REGION Network 8: UnHold Command - controlled by Category Alarm 7
   RUNG wire#powerrail
      Contact( "PackML".Sts.State.Held )
      I_Contact( "UN".Alarm.sts_Category_7_NotLatched )
      Coil( "UN".PackML_Sts_Alarm.cmd_UnHold )
   END_RUNG
   // the same network as SCL:
   "UN".PackML_Sts_Alarm.cmd_UnHold := "PackML".Sts.State.Held AND NOT "UN".Alarm.sts_Category_7_NotLatched;
END_REGION

REGION Network 9: Suspend Command - controlled by Category Alarm 8 or 9
   RUNG wire#powerrail
      Contact( "UN".Alarm.sts_Category_8_NotLatched )
      wire#w1
      Coil( "UN".PackML_Sts_Alarm.cmd_Suspend )
   END_RUNG
   RUNG wire#powerrail
      Contact( "UN".Alarm.sts_Category_9_NotLatched )
   END_RUNG wire#w1
   // the same network as SCL:
   "UN".PackML_Sts_Alarm.cmd_Suspend := "UN".Alarm.sts_Category_8_NotLatched OR "UN".Alarm.sts_Category_9_NotLatched;
END_REGION

REGION Network 10: UnSuspend Command - controlled by clearedCategory Alarm 8 or 9
   RUNG wire#powerrail
      Contact( "PackML".Sts.State.Suspended )
      I_Contact( "UN".Alarm.sts_Category_8_NotLatched )
      I_Contact( "UN".Alarm.sts_Category_9_NotLatched )
      Coil( "UN".PackML_Sts_Alarm.cmd_UnSuspend )
   END_RUNG
   // the same network as SCL:
   "UN".PackML_Sts_Alarm.cmd_UnSuspend := "PackML".Sts.State.Suspended AND NOT "UN".Alarm.sts_Category_8_NotLatched AND NOT "UN".Alarm.sts_Category_9_NotLatched;
END_REGION

REGION Network 11: Clearing SC Command - controlled by clearedCategory Alarm 0 or 1
   RUNG wire#powerrail
      Contact( "PackML".Sts.State.Clearing )
      I_Contact( "UN".Alarm.sts_Category_0_Latched )
      I_Contact( "UN".Alarm.sts_Category_1_Latched )
      Coil( "UN".PackML_Sts_Alarm.sts_Clearing_SC )
   END_RUNG
   // the same network as SCL:
   "UN".PackML_Sts_Alarm.sts_Clearing_SC := "PackML".Sts.State.Clearing AND NOT "UN".Alarm.sts_Category_0_Latched AND NOT "UN".Alarm.sts_Category_1_Latched;
END_REGION

REGION Network 12: Resetting S Command - controlled by clearedCategory Alarm 0-4
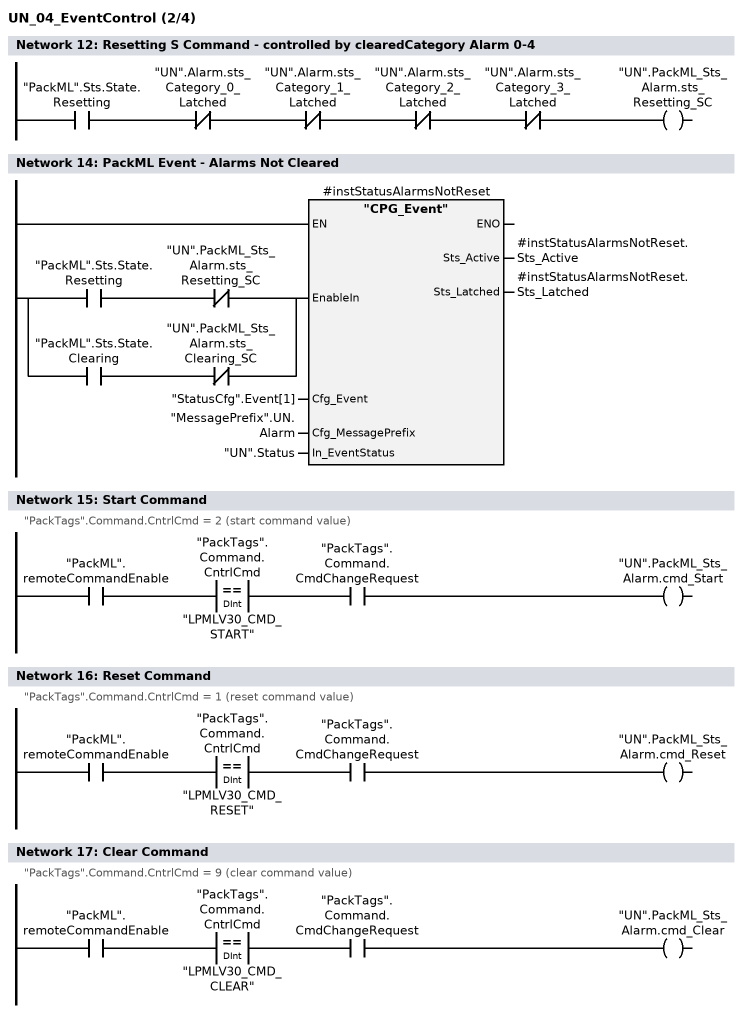
   RUNG wire#powerrail
      Contact( "PackML".Sts.State.Resetting )
      I_Contact( "UN".Alarm.sts_Category_0_Latched )
      I_Contact( "UN".Alarm.sts_Category_1_Latched )
      I_Contact( "UN".Alarm.sts_Category_2_Latched )
      I_Contact( "UN".Alarm.sts_Category_3_Latched )
      Coil( "UN".PackML_Sts_Alarm.sts_Resetting_SC )
   END_RUNG
   // the same network as SCL:
   "UN".PackML_Sts_Alarm.sts_Resetting_SC := "PackML".Sts.State.Resetting AND NOT "UN".Alarm.sts_Category_0_Latched AND NOT "UN".Alarm.sts_Category_1_Latched AND NOT "UN".Alarm.sts_Category_2_Latched AND NOT "UN".Alarm.sts_Category_3_Latched;
END_REGION

REGION Network 13: PackML Event -
END_REGION

REGION Network 14: PackML Event - Alarms Not Cleared
   RUNG wire#powerrail
      #instStatusAlarmsNotReset(EnableIn := wire#w1, Cfg_Event := "StatusCfg".Event[1], Cfg_MessagePrefix := "MessagePrefix".UN.Alarm, In_EventStatus := "UN".Status, Sts_Active => #instStatusAlarmsNotReset.Sts_Active, Sts_Latched => #instStatusAlarmsNotReset.Sts_Latched)
   END_RUNG
   RUNG wire#powerrail
      Contact( "PackML".Sts.State.Resetting )
      I_Contact( "UN".PackML_Sts_Alarm.sts_Resetting_SC )
   END_RUNG wire#w1
   RUNG wire#powerrail
      Contact( "PackML".Sts.State.Clearing )
      I_Contact( "UN".PackML_Sts_Alarm.sts_Clearing_SC )
   END_RUNG wire#w1
   // the same network as SCL:
   #instStatusAlarmsNotReset(EnableIn := ("PackML".Sts.State.Resetting AND NOT "UN".PackML_Sts_Alarm.sts_Resetting_SC) OR ("PackML".Sts.State.Clearing AND NOT "UN".PackML_Sts_Alarm.sts_Clearing_SC),   // "CPG_Event"
                           Cfg_Event := "StatusCfg".Event[1],
                           Cfg_MessagePrefix := "MessagePrefix".UN.Alarm,
                           In_EventStatus := "UN".Status,
                           Sts_Active => #instStatusAlarmsNotReset.Sts_Active,
                           Sts_Latched => #instStatusAlarmsNotReset.Sts_Latched);
END_REGION

REGION Network 15: Start Command
   // "PackTags".Command.CntrlCmd = 2 (start command value)
   RUNG wire#powerrail
      Contact( "PackML".remoteCommandEnable )
      { S7_Templates := "SrcType := DInt" } EQ_Contact(in1 := "PackTags".Command.CntrlCmd, in2 := "LPMLV30_CMD_START")
      Contact( "PackTags".Command.CmdChangeRequest )
      Coil( "UN".PackML_Sts_Alarm.cmd_Start )
   END_RUNG
   // the same network as SCL:
   "UN".PackML_Sts_Alarm.cmd_Start := "PackML".remoteCommandEnable AND ("PackTags".Command.CntrlCmd = "LPMLV30_CMD_START") AND "PackTags".Command.CmdChangeRequest;
END_REGION

REGION Network 16: Reset Command
   // "PackTags".Command.CntrlCmd = 1 (reset command value)
   RUNG wire#powerrail
      Contact( "PackML".remoteCommandEnable )
      { S7_Templates := "SrcType := DInt" } EQ_Contact(in1 := "PackTags".Command.CntrlCmd, in2 := "LPMLV30_CMD_RESET")
      Contact( "PackTags".Command.CmdChangeRequest )
      Coil( "UN".PackML_Sts_Alarm.cmd_Reset )
   END_RUNG
   // the same network as SCL:
   "UN".PackML_Sts_Alarm.cmd_Reset := "PackML".remoteCommandEnable AND ("PackTags".Command.CntrlCmd = "LPMLV30_CMD_RESET") AND "PackTags".Command.CmdChangeRequest;
END_REGION

REGION Network 17: Clear Command
   // "PackTags".Command.CntrlCmd = 9 (clear command value)
   RUNG wire#powerrail
      Contact( "PackML".remoteCommandEnable )
      { S7_Templates := "SrcType := DInt" } EQ_Contact(in1 := "PackTags".Command.CntrlCmd, in2 := "LPMLV30_CMD_CLEAR")
      Contact( "PackTags".Command.CmdChangeRequest )
      Coil( "UN".PackML_Sts_Alarm.cmd_Clear )
   END_RUNG
   // the same network as SCL:
   "UN".PackML_Sts_Alarm.cmd_Clear := "PackML".remoteCommandEnable AND ("PackTags".Command.CntrlCmd = "LPMLV30_CMD_CLEAR") AND "PackTags".Command.CmdChangeRequest;
END_REGION

REGION Network 18: *** EVENT CONTROL MANAGERS ***
END_REGION

REGION Network 19: Reset Command - for all event managers
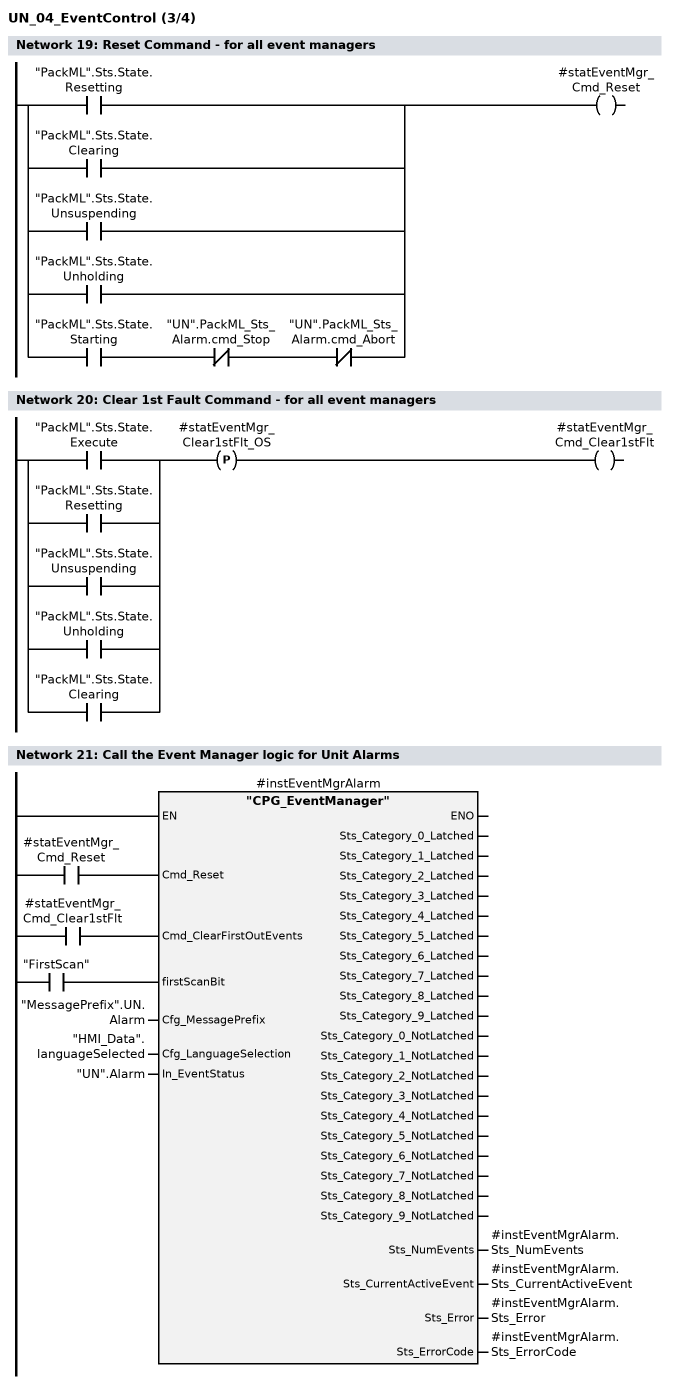
   RUNG wire#powerrail
      Contact( "PackML".Sts.State.Resetting )
      wire#w1
      Coil( #statEventMgr_Cmd_Reset )
   END_RUNG
   RUNG wire#powerrail
      Contact( "PackML".Sts.State.Clearing )
   END_RUNG wire#w1
   RUNG wire#powerrail
      Contact( "PackML".Sts.State.Unsuspending )
   END_RUNG wire#w1
   RUNG wire#powerrail
      Contact( "PackML".Sts.State.Unholding )
   END_RUNG wire#w1
   RUNG wire#powerrail
      Contact( "PackML".Sts.State.Starting )
      I_Contact( "UN".PackML_Sts_Alarm.cmd_Stop )
      I_Contact( "UN".PackML_Sts_Alarm.cmd_Abort )
   END_RUNG wire#w1
   // the same network as SCL:
   #statEventMgr_Cmd_Reset := "PackML".Sts.State.Resetting OR "PackML".Sts.State.Clearing OR "PackML".Sts.State.Unsuspending OR "PackML".Sts.State.Unholding OR ("PackML".Sts.State.Starting AND NOT "UN".PackML_Sts_Alarm.cmd_Stop AND NOT "UN".PackML_Sts_Alarm.cmd_Abort);
END_REGION

REGION Network 20: Clear 1st Fault Command - for all event managers
   RUNG wire#powerrail
      Contact( "PackML".Sts.State.Execute )
      wire#w1
      P_Trig( #statEventMgr_Clear1stFlt_OS )
      Coil( #statEventMgr_Cmd_Clear1stFlt )
   END_RUNG
   RUNG wire#powerrail
      Contact( "PackML".Sts.State.Resetting )
   END_RUNG wire#w1
   RUNG wire#powerrail
      Contact( "PackML".Sts.State.Unsuspending )
   END_RUNG wire#w1
   RUNG wire#powerrail
      Contact( "PackML".Sts.State.Unholding )
   END_RUNG wire#w1
   RUNG wire#powerrail
      Contact( "PackML".Sts.State.Clearing )
   END_RUNG wire#w1
   // the same network as SCL:
   #_w1 := "PackML".Sts.State.Execute OR "PackML".Sts.State.Resetting OR "PackML".Sts.State.Unsuspending OR "PackML".Sts.State.Unholding OR "PackML".Sts.State.Clearing;
   #_w2 := #_w1 AND NOT #statEventMgr_Clear1stFlt_OS;   // rising edge
   #statEventMgr_Clear1stFlt_OS := #_w1;
   #statEventMgr_Cmd_Clear1stFlt := #_w2;
END_REGION

REGION Network 21: Call the Event Manager logic for Unit Alarms
   RUNG wire#powerrail
      #instEventMgrAlarm(Cmd_Reset := wire#w1, Cmd_ClearFirstOutEvents := wire#w2, firstScanBit := wire#w3, Cfg_MessagePrefix := "MessagePrefix".UN.Alarm, Cfg_LanguageSelection := "HMI_Data".languageSelected, In_EventStatus := "UN".Alarm, Sts_Category_0_Latched =>, Sts_Category_1_Latched =>, Sts_Category_2_Latched =>, Sts_Category_3_Latched =>, Sts_Category_4_Latched =>, Sts_Category_5_Latched =>, Sts_Category_6_Latched =>, Sts_Category_7_Latched =>, Sts_Category_8_Latched =>, Sts_Category_9_Latched =>, Sts_Category_0_NotLatched =>, Sts_Category_1_NotLatched =>, Sts_Category_2_NotLatched =>, Sts_Category_3_NotLatched =>, Sts_Category_4_NotLatched =>, Sts_Category_5_NotLatched =>, Sts_Category_6_NotLatched =>, Sts_Category_7_NotLatched =>, Sts_Category_8_NotLatched =>, Sts_Category_9_NotLatched =>, Sts_NumEvents => #instEventMgrAlarm.Sts_NumEvents, Sts_CurrentActiveEvent => #instEventMgrAlarm.Sts_CurrentActiveEvent, Sts_Error => #instEventMgrAlarm.Sts_Error, Sts_ErrorCode => #instEventMgrAlarm.Sts_ErrorCode)
   END_RUNG
   RUNG wire#powerrail
      Contact( #statEventMgr_Cmd_Reset )
   END_RUNG wire#w1
   RUNG wire#powerrail
      Contact( #statEventMgr_Cmd_Clear1stFlt )
   END_RUNG wire#w2
   RUNG wire#powerrail
      Contact( "FirstScan" )
   END_RUNG wire#w3
   // the same network as SCL:
   #instEventMgrAlarm(Cmd_Reset := #statEventMgr_Cmd_Reset,   // "CPG_EventManager"
                      Cmd_ClearFirstOutEvents := #statEventMgr_Cmd_Clear1stFlt,
                      firstScanBit := "FirstScan",
                      Cfg_MessagePrefix := "MessagePrefix".UN.Alarm,
                      Cfg_LanguageSelection := "HMI_Data".languageSelected,
                      In_EventStatus := "UN".Alarm,
                      Sts_NumEvents => #instEventMgrAlarm.Sts_NumEvents,
                      Sts_CurrentActiveEvent => #instEventMgrAlarm.Sts_CurrentActiveEvent,
                      Sts_Error => #instEventMgrAlarm.Sts_Error,
                      Sts_ErrorCode => #instEventMgrAlarm.Sts_ErrorCode);
END_REGION

REGION Network 22: Call the Event Manager logic for Unit Warnings
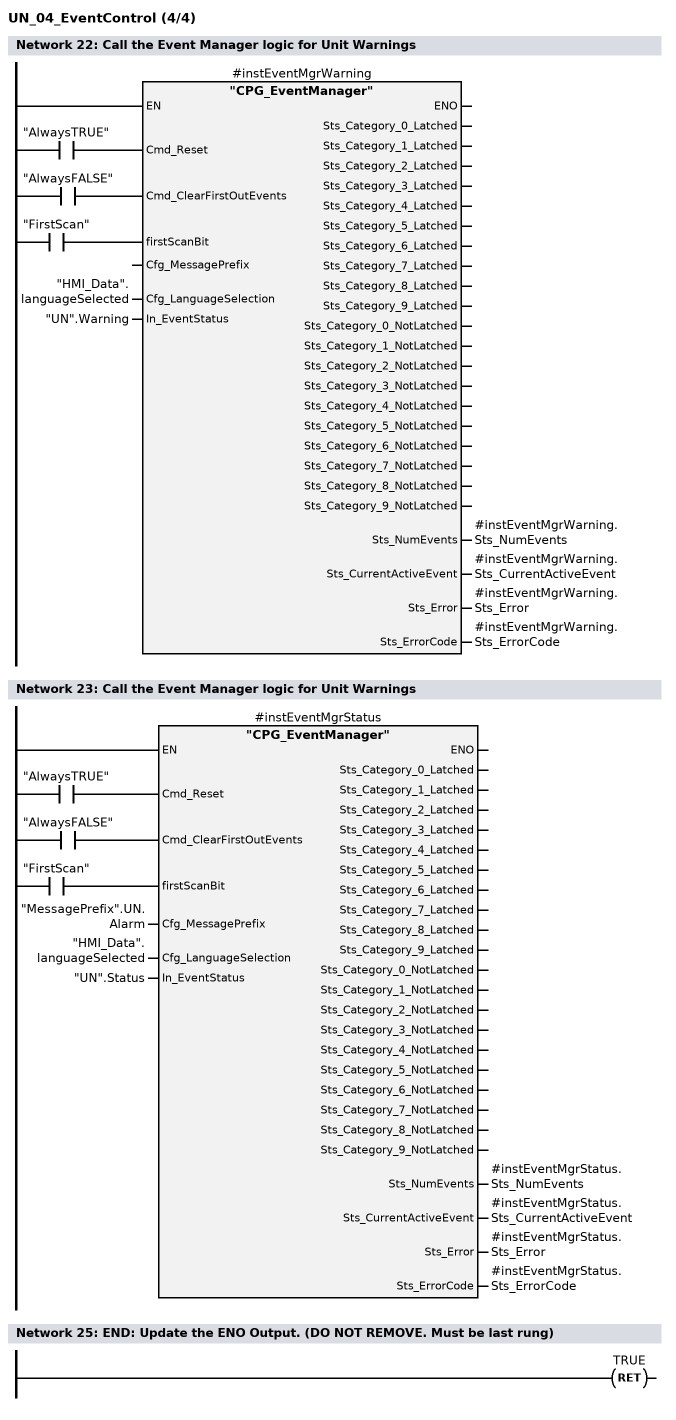
   RUNG wire#powerrail
      #instEventMgrWarning(Cmd_Reset := wire#w1, Cmd_ClearFirstOutEvents := wire#w2, firstScanBit := wire#w3, Cfg_MessagePrefix :=, Cfg_LanguageSelection := "HMI_Data".languageSelected, In_EventStatus := "UN".Warning, Sts_Category_0_Latched =>, Sts_Category_1_Latched =>, Sts_Category_2_Latched =>, Sts_Category_3_Latched =>, Sts_Category_4_Latched =>, Sts_Category_5_Latched =>, Sts_Category_6_Latched =>, Sts_Category_7_Latched =>, Sts_Category_8_Latched =>, Sts_Category_9_Latched =>, Sts_Category_0_NotLatched =>, Sts_Category_1_NotLatched =>, Sts_Category_2_NotLatched =>, Sts_Category_3_NotLatched =>, Sts_Category_4_NotLatched =>, Sts_Category_5_NotLatched =>, Sts_Category_6_NotLatched =>, Sts_Category_7_NotLatched =>, Sts_Category_8_NotLatched =>, Sts_Category_9_NotLatched =>, Sts_NumEvents => #instEventMgrWarning.Sts_NumEvents, Sts_CurrentActiveEvent => #instEventMgrWarning.Sts_CurrentActiveEvent, Sts_Error => #instEventMgrWarning.Sts_Error, Sts_ErrorCode => #instEventMgrWarning.Sts_ErrorCode)
   END_RUNG
   RUNG wire#powerrail
      Contact( "AlwaysTRUE" )
   END_RUNG wire#w1
   RUNG wire#powerrail
      Contact( "AlwaysFALSE" )
   END_RUNG wire#w2
   RUNG wire#powerrail
      Contact( "FirstScan" )
   END_RUNG wire#w3
   // the same network as SCL:
   #instEventMgrWarning(Cmd_Reset := "AlwaysTRUE",   // "CPG_EventManager"
                        Cmd_ClearFirstOutEvents := "AlwaysFALSE",
                        firstScanBit := "FirstScan",
                        Cfg_LanguageSelection := "HMI_Data".languageSelected,
                        In_EventStatus := "UN".Warning,
                        Sts_NumEvents => #instEventMgrWarning.Sts_NumEvents,
                        Sts_CurrentActiveEvent => #instEventMgrWarning.Sts_CurrentActiveEvent,
                        Sts_Error => #instEventMgrWarning.Sts_Error,
                        Sts_ErrorCode => #instEventMgrWarning.Sts_ErrorCode);
END_REGION

REGION Network 23: Call the Event Manager logic for Unit Warnings
   RUNG wire#powerrail
      #instEventMgrStatus(Cmd_Reset := wire#w1, Cmd_ClearFirstOutEvents := wire#w2, firstScanBit := wire#w3, Cfg_MessagePrefix := "MessagePrefix".UN.Alarm, Cfg_LanguageSelection := "HMI_Data".languageSelected, In_EventStatus := "UN".Status, Sts_Category_0_Latched =>, Sts_Category_1_Latched =>, Sts_Category_2_Latched =>, Sts_Category_3_Latched =>, Sts_Category_4_Latched =>, Sts_Category_5_Latched =>, Sts_Category_6_Latched =>, Sts_Category_7_Latched =>, Sts_Category_8_Latched =>, Sts_Category_9_Latched =>, Sts_Category_0_NotLatched =>, Sts_Category_1_NotLatched =>, Sts_Category_2_NotLatched =>, Sts_Category_3_NotLatched =>, Sts_Category_4_NotLatched =>, Sts_Category_5_NotLatched =>, Sts_Category_6_NotLatched =>, Sts_Category_7_NotLatched =>, Sts_Category_8_NotLatched =>, Sts_Category_9_NotLatched =>, Sts_NumEvents => #instEventMgrStatus.Sts_NumEvents, Sts_CurrentActiveEvent => #instEventMgrStatus.Sts_CurrentActiveEvent, Sts_Error => #instEventMgrStatus.Sts_Error, Sts_ErrorCode => #instEventMgrStatus.Sts_ErrorCode)
   END_RUNG
   RUNG wire#powerrail
      Contact( "AlwaysTRUE" )
   END_RUNG wire#w1
   RUNG wire#powerrail
      Contact( "AlwaysFALSE" )
   END_RUNG wire#w2
   RUNG wire#powerrail
      Contact( "FirstScan" )
   END_RUNG wire#w3
   // the same network as SCL:
   #instEventMgrStatus(Cmd_Reset := "AlwaysTRUE",   // "CPG_EventManager"
                       Cmd_ClearFirstOutEvents := "AlwaysFALSE",
                       firstScanBit := "FirstScan",
                       Cfg_MessagePrefix := "MessagePrefix".UN.Alarm,
                       Cfg_LanguageSelection := "HMI_Data".languageSelected,
                       In_EventStatus := "UN".Status,
                       Sts_NumEvents => #instEventMgrStatus.Sts_NumEvents,
                       Sts_CurrentActiveEvent => #instEventMgrStatus.Sts_CurrentActiveEvent,
                       Sts_Error => #instEventMgrStatus.Sts_Error,
                       Sts_ErrorCode => #instEventMgrStatus.Sts_ErrorCode);
END_REGION

REGION Network 25: END: Update the ENO Output. (DO NOT REMOVE. Must be last rung)
   RUNG wire#powerrail
      ReturnCoil( TRUE )
   END_RUNG
   // the same network as SCL:
   ENO := TRUE;
   RETURN;
END_REGION
END_FUNCTION_BLOCK

FUNCTION_BLOCK "UN_05_EventSummation"   // FB31625, LAD
TITLE = UN_05_EventSummation
{ S7_Optimized_Access := 'TRUE' }
AUTHOR : tech.team.motioncontrol@siemens.com
FAMILY : CPG
VERSION : 1.1
// Support: tech.team.motioncontrol@siemens.com
   VAR
      instEventSumBeg_Alarm : "CPG_EventSummationBegin";   // instanceFB - EventSummationBegin - Alarm Events
      instEventSum_Alarm_UN : "CPG_EventSummation";   // instanceFB - EventSummation FB - Alarm Events - UN
      instEventSum_Alarm_EM00 : "CPG_EventSummation";   // instanceFB - EventSummation FB - Alarm Events - EM00
      instEventSum_Alarm_EM01 : "CPG_EventSummation";   // instanceFB - EventSummation FB - Alarm Events - EM01
      instEventSum_Alarm_EM02 : "CPG_EventSummation";   // instanceFB - EventSummation FB - Alarm Events - EM02
      instEventSumEnd_Alarm : "CPG_EventSummationEnd";   // instanceFB - EventSummationEnd - Alarm Events
      instEventSortFilter_Alarm : "CPG_EventSortFilter";   // instanceFB - EventSortFilter FB - Alarms
      instAlarmMove : "CPG_AlarmMove";   // instance FB - Alarm Move
      instEventSumBeg_Warning : "CPG_EventSummationBegin";   // instanceFB - EventSummationBegin - Warning Events
      instEventSum_Warning_UN : "CPG_EventSummation";   // instanceFB - EventSummation FB - Warning Events - UN
      instEventSum_Warning_EM00 : "CPG_EventSummation";   // instanceFB - EventSummation FB - Warning Events - EM00
      instEventSum_Warning_EM01 : "CPG_EventSummation";   // instanceFB - EventSummation FB - Warning Events - EM01
      instEventSum_Warning_EM02 : "CPG_EventSummation";   // instanceFB - EventSummation FB - Warning Events - EM02
      instEventSumEnd_Warning : "CPG_EventSummationEnd";   // instanceFB - EventSummationEnd - Warning Events
      instEventSortFilter_Warning : "CPG_EventSortFilter";   // instanceFB - EventSortFilter FB - Alarms
      instWarning_MsgScroll : "CPG_MsgScroll";   // instance FB - Warning Scroll
      instEventSumBeg_Status : "CPG_EventSummationBegin";   // instanceFB - EventSummationBegin - Status Events
      instEventSum_Status_UN : "CPG_EventSummation";   // instanceFB - EventSummation FB - Status Events - UN
      instEventSum_Status_EM00 : "CPG_EventSummation";   // instanceFB - EventSummation FB - Status Events - EM00
      instEventSum_Status_EM01 : "CPG_EventSummation";   // instanceFB - EventSummation FB - Status Events - EM01
      instEventSum_Status_EM02 : "CPG_EventSummation";   // instanceFB - EventSummation FB - Status Events - EM02
      instEventSumEnd_Status : "CPG_EventSummationEnd";   // instanceFB - EventSummationEnd - Status Events
      instPackML_AlarmHistory : "CPG_AlarmHistory";   // instance FB - Capturing the 1st fault history
      instProgram_Alarm : Program_Alarm;   // instance DB for Program Alarm - diag to PLC HMI
      instWarningMove : "CPG_AlarmMove";
      instPareto : "CPG_ParetoAnalysis";
   END_VAR
   VAR_TEMP
      tempAlarmMove_Sts_Error : Bool;   // Error with AlarmMove?
      tempAlarmMove_Sts_ErrorCode : Int;   // AlarmMove Error code
      tempProgramAlarm_error : Bool;
      tempProgramAlarm_status : Word;
   END_VAR
BEGIN

REGION Network 1: Call the Alarm Event Summary - Beginning FB
   // **********  ALARM CONTROL SUMMATION  **********
   //  
   // The event summation begin instruction prepares the summation blocks.  It should 
   // be run each time before the FB_EventSummation blocks.
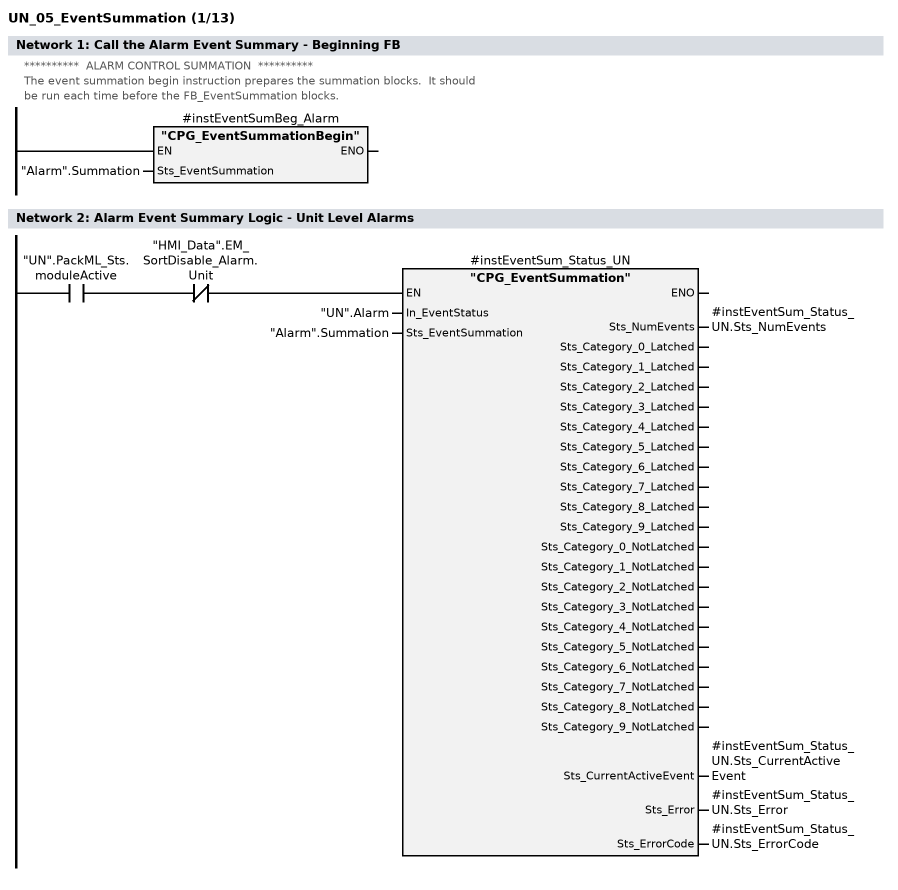
   RUNG wire#powerrail
      #instEventSumBeg_Alarm(Sts_EventSummation := "Alarm".Summation)
   END_RUNG
   // the same network as SCL:
   #instEventSumBeg_Alarm(Sts_EventSummation := "Alarm".Summation);   // "CPG_EventSummationBegin"
END_REGION

REGION Network 2: Alarm Event Summary Logic - Unit Level Alarms
   RUNG wire#powerrail
      Contact( "UN".PackML_Sts.moduleActive )
      I_Contact( "HMI_Data".EM_SortDisable_Alarm.Unit )
      #instEventSum_Status_UN(In_EventStatus := "UN".Alarm, Sts_EventSummation := "Alarm".Summation, Sts_NumEvents => #instEventSum_Status_UN.Sts_NumEvents, Sts_Category_0_Latched =>, Sts_Category_1_Latched =>, Sts_Category_2_Latched =>, Sts_Category_3_Latched =>, Sts_Category_4_Latched =>, Sts_Category_5_Latched =>, Sts_Category_6_Latched =>, Sts_Category_7_Latched =>, Sts_Category_8_Latched =>, Sts_Category_9_Latched =>, Sts_Category_0_NotLatched =>, Sts_Category_1_NotLatched =>, Sts_Category_2_NotLatched =>, Sts_Category_3_NotLatched =>, Sts_Category_4_NotLatched =>, Sts_Category_5_NotLatched =>, Sts_Category_6_NotLatched =>, Sts_Category_7_NotLatched =>, Sts_Category_8_NotLatched =>, Sts_Category_9_NotLatched =>, Sts_CurrentActiveEvent => #instEventSum_Status_UN.Sts_CurrentActiveEvent, Sts_Error => #instEventSum_Status_UN.Sts_Error, Sts_ErrorCode => #instEventSum_Status_UN.Sts_ErrorCode)
   END_RUNG
   // the same network as SCL:
   IF "UN".PackML_Sts.moduleActive AND NOT "HMI_Data".EM_SortDisable_Alarm.Unit THEN
       #instEventSum_Status_UN(In_EventStatus := "UN".Alarm,   // "CPG_EventSummation"
                               Sts_EventSummation := "Alarm".Summation,
                               Sts_NumEvents => #instEventSum_Status_UN.Sts_NumEvents,
                               Sts_CurrentActiveEvent => #instEventSum_Status_UN.Sts_CurrentActiveEvent,
                               Sts_Error => #instEventSum_Status_UN.Sts_Error,
                               Sts_ErrorCode => #instEventSum_Status_UN.Sts_ErrorCode);
   END_IF;
END_REGION

REGION Network 3: Alarm Event Summary Logic - Equipment Module #00
   // This instance of the Event Sum (or Event Summation) is used to merge the events 
   // from EM0 into the larger Unit or UN evevts list.
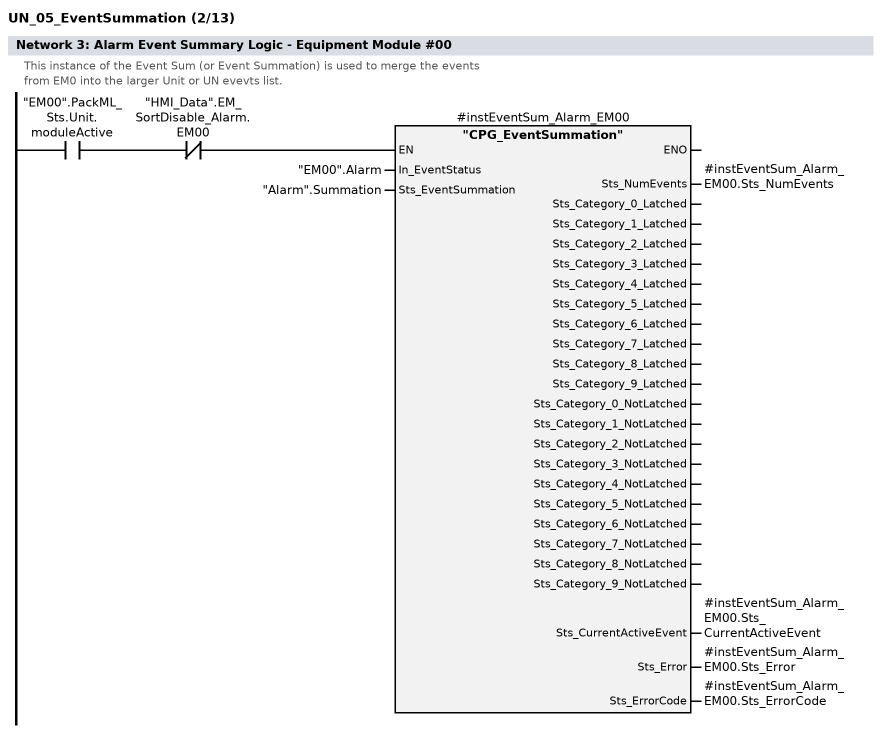
   RUNG wire#powerrail
      Contact( "EM00".PackML_Sts.Unit.moduleActive )
      I_Contact( "HMI_Data".EM_SortDisable_Alarm.EM00 )
      #instEventSum_Alarm_EM00(In_EventStatus := "EM00".Alarm, Sts_EventSummation := "Alarm".Summation, Sts_NumEvents => #instEventSum_Alarm_EM00.Sts_NumEvents, Sts_Category_0_Latched =>, Sts_Category_1_Latched =>, Sts_Category_2_Latched =>, Sts_Category_3_Latched =>, Sts_Category_4_Latched =>, Sts_Category_5_Latched =>, Sts_Category_6_Latched =>, Sts_Category_7_Latched =>, Sts_Category_8_Latched =>, Sts_Category_9_Latched =>, Sts_Category_0_NotLatched =>, Sts_Category_1_NotLatched =>, Sts_Category_2_NotLatched =>, Sts_Category_3_NotLatched =>, Sts_Category_4_NotLatched =>, Sts_Category_5_NotLatched =>, Sts_Category_6_NotLatched =>, Sts_Category_7_NotLatched =>, Sts_Category_8_NotLatched =>, Sts_Category_9_NotLatched =>, Sts_CurrentActiveEvent => #instEventSum_Alarm_EM00.Sts_CurrentActiveEvent, Sts_Error => #instEventSum_Alarm_EM00.Sts_Error, Sts_ErrorCode => #instEventSum_Alarm_EM00.Sts_ErrorCode)
   END_RUNG
   // the same network as SCL:
   IF "EM00".PackML_Sts.Unit.moduleActive AND NOT "HMI_Data".EM_SortDisable_Alarm.EM00 THEN
       #instEventSum_Alarm_EM00(In_EventStatus := "EM00".Alarm,   // "CPG_EventSummation"
                               Sts_EventSummation := "Alarm".Summation,
                               Sts_NumEvents => #instEventSum_Alarm_EM00.Sts_NumEvents,
                               Sts_CurrentActiveEvent => #instEventSum_Alarm_EM00.Sts_CurrentActiveEvent,
                               Sts_Error => #instEventSum_Alarm_EM00.Sts_Error,
                               Sts_ErrorCode => #instEventSum_Alarm_EM00.Sts_ErrorCode);
   END_IF;
END_REGION

REGION Network 4: Alarm Event Summary Logic - Equipment Module #01
   // This instance of the Event Sum (or Event Summation) is used to merge the events 
   // from EM01 into the larger Unit or UN evevts list.
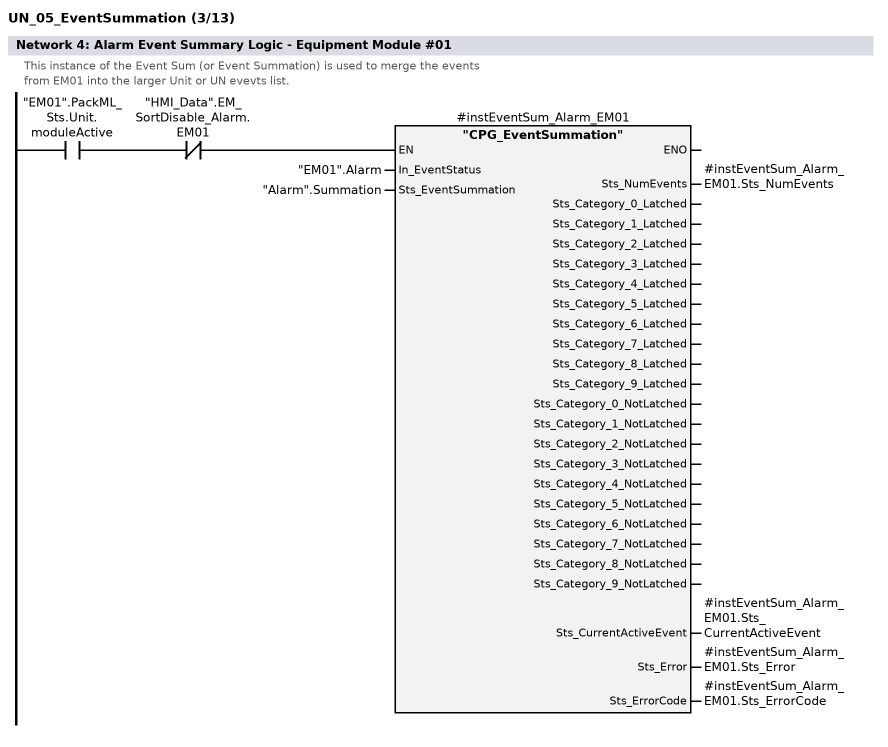
   RUNG wire#powerrail
      Contact( "EM01".PackML_Sts.Unit.moduleActive )
      I_Contact( "HMI_Data".EM_SortDisable_Alarm.EM01 )
      #instEventSum_Alarm_EM01(In_EventStatus := "EM01".Alarm, Sts_EventSummation := "Alarm".Summation, Sts_NumEvents => #instEventSum_Alarm_EM01.Sts_NumEvents, Sts_Category_0_Latched =>, Sts_Category_1_Latched =>, Sts_Category_2_Latched =>, Sts_Category_3_Latched =>, Sts_Category_4_Latched =>, Sts_Category_5_Latched =>, Sts_Category_6_Latched =>, Sts_Category_7_Latched =>, Sts_Category_8_Latched =>, Sts_Category_9_Latched =>, Sts_Category_0_NotLatched =>, Sts_Category_1_NotLatched =>, Sts_Category_2_NotLatched =>, Sts_Category_3_NotLatched =>, Sts_Category_4_NotLatched =>, Sts_Category_5_NotLatched =>, Sts_Category_6_NotLatched =>, Sts_Category_7_NotLatched =>, Sts_Category_8_NotLatched =>, Sts_Category_9_NotLatched =>, Sts_CurrentActiveEvent => #instEventSum_Alarm_EM01.Sts_CurrentActiveEvent, Sts_Error => #instEventSum_Alarm_EM01.Sts_Error, Sts_ErrorCode => #instEventSum_Alarm_EM01.Sts_ErrorCode)
   END_RUNG
   // the same network as SCL:
   IF "EM01".PackML_Sts.Unit.moduleActive AND NOT "HMI_Data".EM_SortDisable_Alarm.EM01 THEN
       #instEventSum_Alarm_EM01(In_EventStatus := "EM01".Alarm,   // "CPG_EventSummation"
                               Sts_EventSummation := "Alarm".Summation,
                               Sts_NumEvents => #instEventSum_Alarm_EM01.Sts_NumEvents,
                               Sts_CurrentActiveEvent => #instEventSum_Alarm_EM01.Sts_CurrentActiveEvent,
                               Sts_Error => #instEventSum_Alarm_EM01.Sts_Error,
                               Sts_ErrorCode => #instEventSum_Alarm_EM01.Sts_ErrorCode);
   END_IF;
END_REGION

REGION Network 5: Alarm Event Summary Logic - Equipment Module #02
   // This instance of the Event Sum (or Event Summation) is used to merge the events 
   // from EM01 into the larger Unit or UN evevts list.
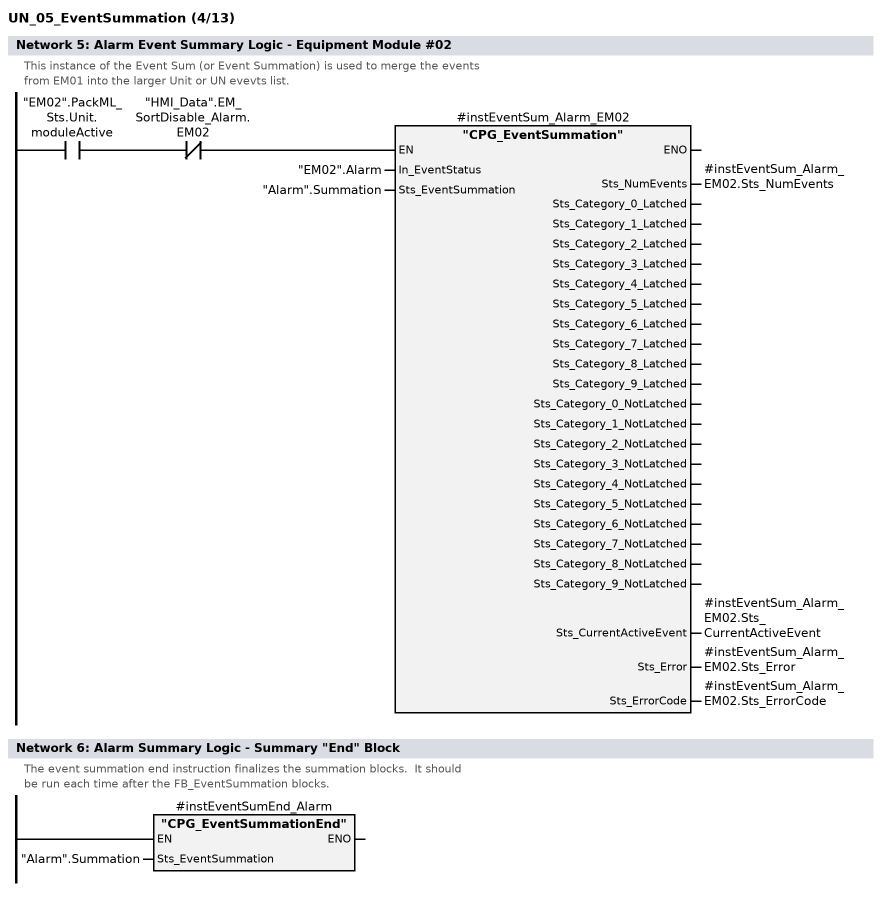
   RUNG wire#powerrail
      Contact( "EM02".PackML_Sts.Unit.moduleActive )
      I_Contact( "HMI_Data".EM_SortDisable_Alarm.EM02 )
      #instEventSum_Alarm_EM02(In_EventStatus := "EM02".Alarm, Sts_EventSummation := "Alarm".Summation, Sts_NumEvents => #instEventSum_Alarm_EM02.Sts_NumEvents, Sts_Category_0_Latched =>, Sts_Category_1_Latched =>, Sts_Category_2_Latched =>, Sts_Category_3_Latched =>, Sts_Category_4_Latched =>, Sts_Category_5_Latched =>, Sts_Category_6_Latched =>, Sts_Category_7_Latched =>, Sts_Category_8_Latched =>, Sts_Category_9_Latched =>, Sts_Category_0_NotLatched =>, Sts_Category_1_NotLatched =>, Sts_Category_2_NotLatched =>, Sts_Category_3_NotLatched =>, Sts_Category_4_NotLatched =>, Sts_Category_5_NotLatched =>, Sts_Category_6_NotLatched =>, Sts_Category_7_NotLatched =>, Sts_Category_8_NotLatched =>, Sts_Category_9_NotLatched =>, Sts_CurrentActiveEvent => #instEventSum_Alarm_EM02.Sts_CurrentActiveEvent, Sts_Error => #instEventSum_Alarm_EM02.Sts_Error, Sts_ErrorCode => #instEventSum_Alarm_EM02.Sts_ErrorCode)
   END_RUNG
   // the same network as SCL:
   IF "EM02".PackML_Sts.Unit.moduleActive AND NOT "HMI_Data".EM_SortDisable_Alarm.EM02 THEN
       #instEventSum_Alarm_EM02(In_EventStatus := "EM02".Alarm,   // "CPG_EventSummation"
                               Sts_EventSummation := "Alarm".Summation,
                               Sts_NumEvents => #instEventSum_Alarm_EM02.Sts_NumEvents,
                               Sts_CurrentActiveEvent => #instEventSum_Alarm_EM02.Sts_CurrentActiveEvent,
                               Sts_Error => #instEventSum_Alarm_EM02.Sts_Error,
                               Sts_ErrorCode => #instEventSum_Alarm_EM02.Sts_ErrorCode);
   END_IF;
END_REGION

REGION Network 6: Alarm Summary Logic - Summary "End" Block
   // The event summation end instruction finalizes the summation blocks.  It should 
   // be run each time after the FB_EventSummation blocks.
   RUNG wire#powerrail
      #instEventSumEnd_Alarm(Sts_EventSummation := "Alarm".Summation)
   END_RUNG
   // the same network as SCL:
   #instEventSumEnd_Alarm(Sts_EventSummation := "Alarm".Summation);   // "CPG_EventSummationEnd"
END_REGION

REGION Network 7: Update Admin.Alarm information.
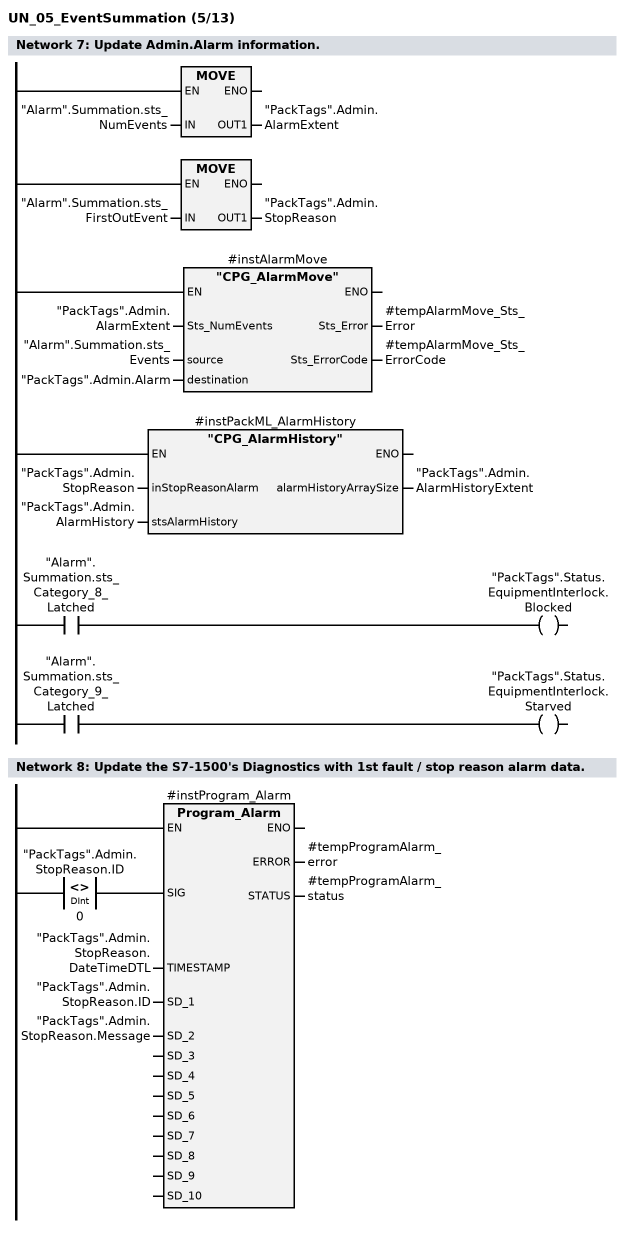
   RUNG wire#powerrail
      { S7_GenerateENO := "TRUE" } Move(in := "Alarm".Summation.sts_NumEvents, out1 => "PackTags".Admin.AlarmExtent)
   END_RUNG
   RUNG wire#powerrail
      Move(in := "Alarm".Summation.sts_FirstOutEvent, out1 => "PackTags".Admin.StopReason)
   END_RUNG
   RUNG wire#powerrail
      #instAlarmMove(Sts_NumEvents := "PackTags".Admin.AlarmExtent, source := "Alarm".Summation.sts_Events, destination := "PackTags".Admin.Alarm, Sts_Error => #tempAlarmMove_Sts_Error, Sts_ErrorCode => #tempAlarmMove_Sts_ErrorCode)
   END_RUNG
   RUNG wire#powerrail
      #instPackML_AlarmHistory(inStopReasonAlarm := "PackTags".Admin.StopReason, stsAlarmHistory := "PackTags".Admin.AlarmHistory, alarmHistoryArraySize => "PackTags".Admin.AlarmHistoryExtent)
   END_RUNG
   RUNG wire#powerrail
      Contact( "Alarm".Summation.sts_Category_8_Latched )
      Coil( "PackTags".Status.EquipmentInterlock.Blocked )
   END_RUNG
   RUNG wire#powerrail
      Contact( "Alarm".Summation.sts_Category_9_Latched )
      Coil( "PackTags".Status.EquipmentInterlock.Starved )
   END_RUNG
   // the same network as SCL:
   "PackTags".Admin.AlarmExtent := "Alarm".Summation.sts_NumEvents;
   "PackTags".Admin.StopReason := "Alarm".Summation.sts_FirstOutEvent;
   #instAlarmMove(Sts_NumEvents := "PackTags".Admin.AlarmExtent,   // "CPG_AlarmMove"
                  source := "Alarm".Summation.sts_Events,
                  destination := "PackTags".Admin.Alarm,
                  Sts_Error => #tempAlarmMove_Sts_Error,
                  Sts_ErrorCode => #tempAlarmMove_Sts_ErrorCode);
   #instPackML_AlarmHistory(inStopReasonAlarm := "PackTags".Admin.StopReason,   // "CPG_AlarmHistory"
                           stsAlarmHistory := "PackTags".Admin.AlarmHistory,
                           alarmHistoryArraySize => "PackTags".Admin.AlarmHistoryExtent);
   "PackTags".Status.EquipmentInterlock.Blocked := "Alarm".Summation.sts_Category_8_Latched;
   "PackTags".Status.EquipmentInterlock.Starved := "Alarm".Summation.sts_Category_9_Latched;
END_REGION

REGION Network 8: Update the S7-1500's Diagnostics with 1st fault / stop reason alarm data.
   #instProgram_Alarm(SIG := "PackTags".Admin.StopReason.ID <> 0,   // Program_Alarm
                      TIMESTAMP := "PackTags".Admin.StopReason.DateTimeDTL,
                      SD_1 := "PackTags".Admin.StopReason.ID,
                      SD_2 := "PackTags".Admin.StopReason.Message,
                      Error => #tempProgramAlarm_error,
                      Status => #tempProgramAlarm_status);
END_REGION

REGION Network 9: Event Sort Filter logic - Alarms
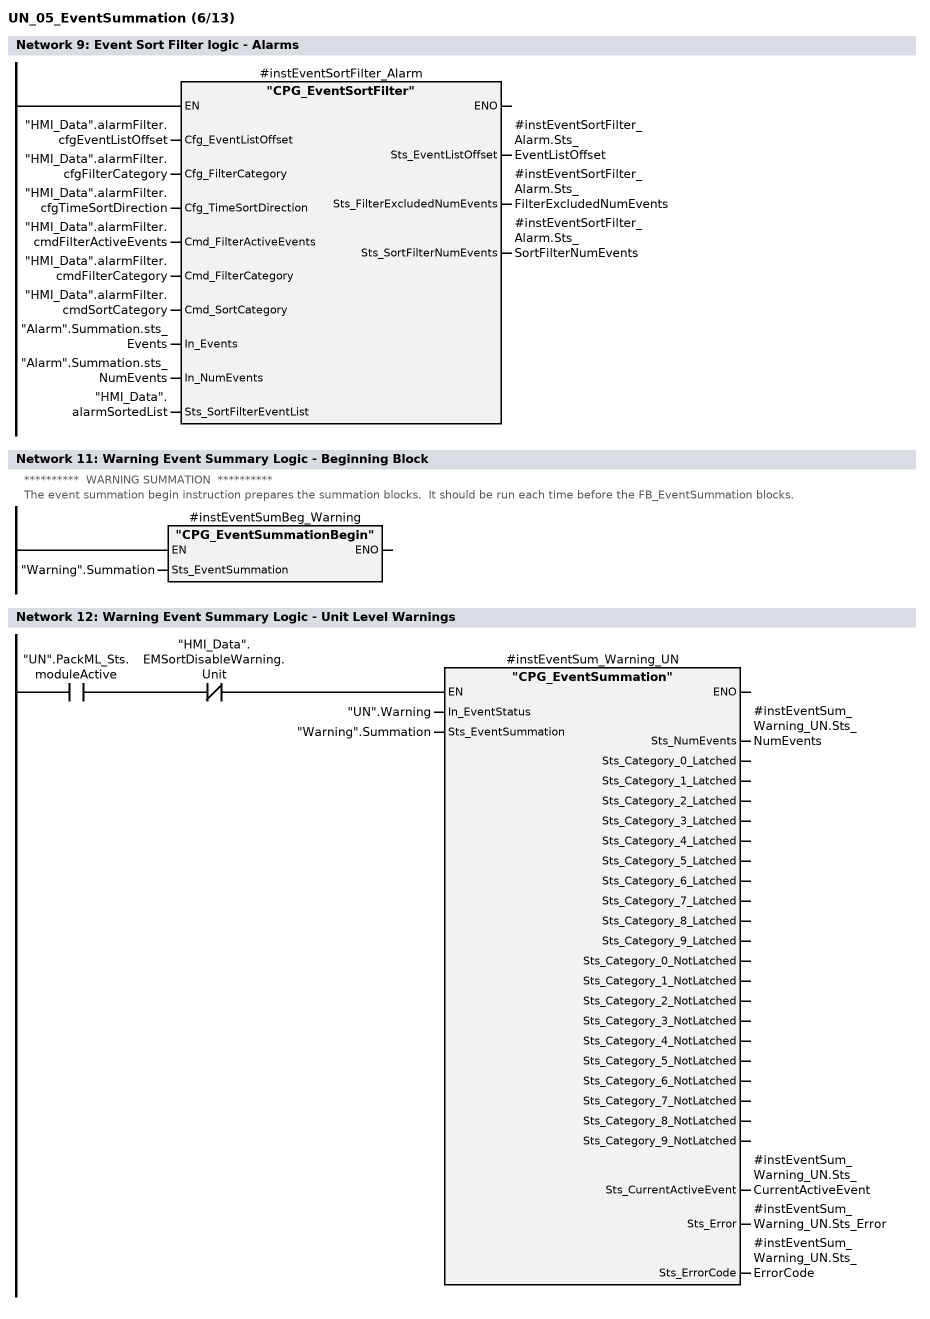
   RUNG wire#powerrail
      #instEventSortFilter_Alarm(Cfg_EventListOffset := "HMI_Data".alarmFilter.cfgEventListOffset, Cfg_FilterCategory := "HMI_Data".alarmFilter.cfgFilterCategory, Cfg_TimeSortDirection := "HMI_Data".alarmFilter.cfgTimeSortDirection, Cmd_FilterActiveEvents := "HMI_Data".alarmFilter.cmdFilterActiveEvents, Cmd_FilterCategory := "HMI_Data".alarmFilter.cmdFilterCategory, Cmd_SortCategory := "HMI_Data".alarmFilter.cmdSortCategory, In_Events := "Alarm".Summation.sts_Events, In_NumEvents := "Alarm".Summation.sts_NumEvents, Sts_SortFilterEventList := "HMI_Data".alarmSortedList, Sts_EventListOffset => #instEventSortFilter_Alarm.Sts_EventListOffset, Sts_FilterExcludedNumEvents => #instEventSortFilter_Alarm.Sts_FilterExcludedNumEvents, Sts_SortFilterNumEvents => #instEventSortFilter_Alarm.Sts_SortFilterNumEvents)
   END_RUNG
   // the same network as SCL:
   #instEventSortFilter_Alarm(Cfg_EventListOffset := "HMI_Data".alarmFilter.cfgEventListOffset,   // "CPG_EventSortFilter"
                           Cfg_FilterCategory := "HMI_Data".alarmFilter.cfgFilterCategory,
                           Cfg_TimeSortDirection := "HMI_Data".alarmFilter.cfgTimeSortDirection,
                           Cmd_FilterActiveEvents := "HMI_Data".alarmFilter.cmdFilterActiveEvents,
                           Cmd_FilterCategory := "HMI_Data".alarmFilter.cmdFilterCategory,
                           Cmd_SortCategory := "HMI_Data".alarmFilter.cmdSortCategory,
                           In_Events := "Alarm".Summation.sts_Events,
                           In_NumEvents := "Alarm".Summation.sts_NumEvents,
                           Sts_SortFilterEventList := "HMI_Data".alarmSortedList,
                           Sts_EventListOffset => #instEventSortFilter_Alarm.Sts_EventListOffset,